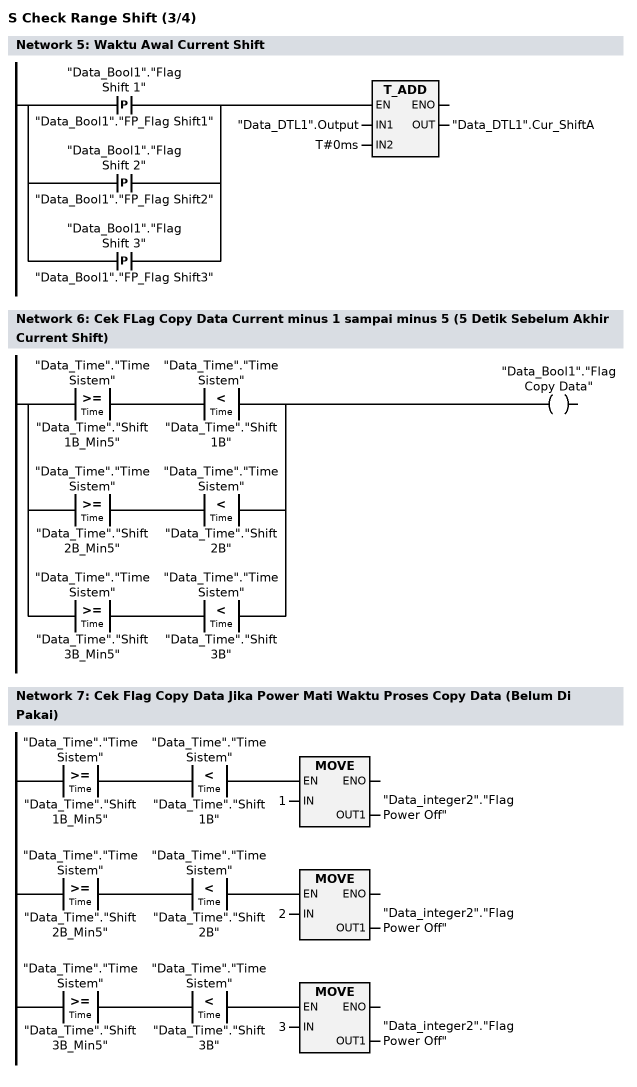
   #_w1 := "Data_Bool1"."Flag Shift 1" AND NOT "Data_Bool1"."FP_Flag Shift1";   // rising edge of "Data_Bool1"."Flag Shift 1"
   "Data_Bool1"."FP_Flag Shift1" := "Data_Bool1"."Flag Shift 1";
   #_w2 := "Data_Bool1"."Flag Shift 2" AND NOT "Data_Bool1"."FP_Flag Shift2";   // rising edge of "Data_Bool1"."Flag Shift 2"
   "Data_Bool1"."FP_Flag Shift2" := "Data_Bool1"."Flag Shift 2";
   #_w3 := "Data_Bool1"."Flag Shift 3" AND NOT "Data_Bool1"."FP_Flag Shift3";   // rising edge of "Data_Bool1"."Flag Shift 3"
   "Data_Bool1"."FP_Flag Shift3" := "Data_Bool1"."Flag Shift 3";
   IF #_w1 OR #_w2 OR #_w3 THEN
       "Data_DTL1".Cur_ShiftA := T_ADD(IN1 := "Data_DTL1".Output, IN2 := T#0ms);
   END_IF;
END_REGION

REGION Network 6: Cek FLag Copy Data Current minus 1 sampai minus 5 (5 Detik Sebelum Akhir Current Shift)
   RUNG wire#powerrail
      { S7_Templates := "SrcType := Time" } GE_Contact(in1 := "Data_Time"."Time Sistem", in2 := "Data_Time"."Shift 1B_Min5")
      { S7_Templates := "SrcType := Time" } LT_Contact(in1 := "Data_Time"."Time Sistem", in2 := "Data_Time"."Shift 1B")
      wire#w1
      Coil( "Data_Bool1"."Flag Copy Data" )
   END_RUNG
   RUNG wire#powerrail
      { S7_Templates := "SrcType := Time" } GE_Contact(in1 := "Data_Time"."Time Sistem", in2 := "Data_Time"."Shift 2B_Min5")
      { S7_Templates := "SrcType := Time" } LT_Contact(in1 := "Data_Time"."Time Sistem", in2 := "Data_Time"."Shift 2B")
   END_RUNG wire#w1
   RUNG wire#powerrail
      { S7_Templates := "SrcType := Time" } GE_Contact(in1 := "Data_Time"."Time Sistem", in2 := "Data_Time"."Shift 3B_Min5")
      { S7_Templates := "SrcType := Time" } LT_Contact(in1 := "Data_Time"."Time Sistem", in2 := "Data_Time"."Shift 3B")
   END_RUNG wire#w1
   // the same network as SCL:
   "Data_Bool1"."Flag Copy Data" := (("Data_Time"."Time Sistem" >= "Data_Time"."Shift 1B_Min5") AND ("Data_Time"."Time Sistem" < "Data_Time"."Shift 1B")) OR (("Data_Time"."Time Sistem" >= "Data_Time"."Shift 2B_Min5") AND ("Data_Time"."Time Sistem" < "Data_Time"."Shift 2B")) OR (("Data_Time"."Time Sistem" >= "Data_Time"."Shift 3B_Min5") AND ("Data_Time"."Time Sistem" < "Data_Time"."Shift 3B"));
END_REGION

REGION Network 7: Cek Flag Copy Data Jika Power Mati Waktu Proses Copy Data (Belum Di Pakai)
   RUNG wire#powerrail
      { S7_Templates := "SrcType := Time" } GE_Contact(in1 := "Data_Time"."Time Sistem", in2 := "Data_Time"."Shift 1B_Min5")
      { S7_Templates := "SrcType := Time" } LT_Contact(in1 := "Data_Time"."Time Sistem", in2 := "Data_Time"."Shift 1B")
      { S7_GenerateENO := "TRUE" } Move(in := 1, out1 => "Data_integer2"."Flag Power Off")
   END_RUNG
   RUNG wire#powerrail
      { S7_Templates := "SrcType := Time" } GE_Contact(in1 := "Data_Time"."Time Sistem", in2 := "Data_Time"."Shift 2B_Min5")
      { S7_Templates := "SrcType := Time" } LT_Contact(in1 := "Data_Time"."Time Sistem", in2 := "Data_Time"."Shift 2B")
      { S7_GenerateENO := "TRUE" } Move(in := 2, out1 => "Data_integer2"."Flag Power Off")
   END_RUNG
   RUNG wire#powerrail
      { S7_Templates := "SrcType := Time" } GE_Contact(in1 := "Data_Time"."Time Sistem", in2 := "Data_Time"."Shift 3B_Min5")
      { S7_Templates := "SrcType := Time" } LT_Contact(in1 := "Data_Time"."Time Sistem", in2 := "Data_Time"."Shift 3B")
      { S7_GenerateENO := "TRUE" } Move(in := 3, out1 => "Data_integer2"."Flag Power Off")
   END_RUNG
   // the same network as SCL:
   IF ("Data_Time"."Time Sistem" >= "Data_Time"."Shift 1B_Min5") AND ("Data_Time"."Time Sistem" < "Data_Time"."Shift 1B") THEN
       "Data_integer2"."Flag Power Off" := 1;
   END_IF;
   IF ("Data_Time"."Time Sistem" >= "Data_Time"."Shift 2B_Min5") AND ("Data_Time"."Time Sistem" < "Data_Time"."Shift 2B") THEN
       "Data_integer2"."Flag Power Off" := 2;
   END_IF;
   IF ("Data_Time"."Time Sistem" >= "Data_Time"."Shift 3B_Min5") AND ("Data_Time"."Time Sistem" < "Data_Time"."Shift 3B") THEN
       "Data_integer2"."Flag Power Off" := 3;
   END_IF;
END_REGION

REGION Network 8: Waktu Awal Current Shift Static Dan Set Copi data Setelah Power mati di waktu proses Copi Data (belum Dipakai)
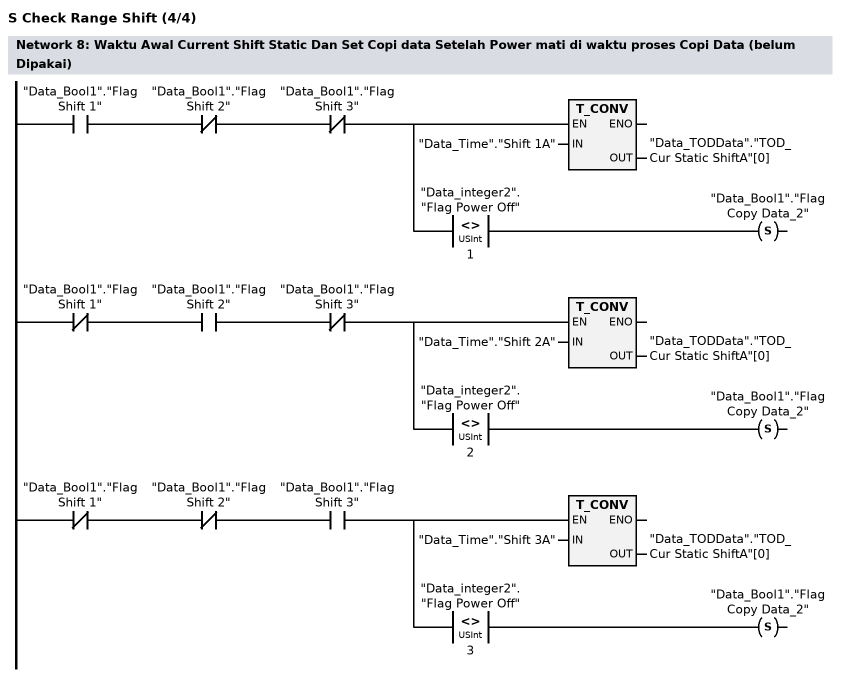
   #_w1 := "Data_Bool1"."Flag Shift 1" AND NOT "Data_Bool1"."Flag Shift 2" AND NOT "Data_Bool1"."Flag Shift 3";
   IF #_w1 THEN "Data_TODData"."TOD_Cur Static ShiftA"[0] := T_CONV(IN := "Data_Time"."Shift 1A"); END_IF;
   IF #_w1 AND ("Data_integer2"."Flag Power Off" <> 1) THEN "Data_Bool1"."Flag Copy Data_2" := TRUE; END_IF;
   #_w2 := NOT "Data_Bool1"."Flag Shift 1" AND "Data_Bool1"."Flag Shift 2" AND NOT "Data_Bool1"."Flag Shift 3";
   IF #_w2 THEN "Data_TODData"."TOD_Cur Static ShiftA"[0] := T_CONV(IN := "Data_Time"."Shift 2A"); END_IF;
   IF #_w2 AND ("Data_integer2"."Flag Power Off" <> 2) THEN "Data_Bool1"."Flag Copy Data_2" := TRUE; END_IF;
   #_w3 := NOT "Data_Bool1"."Flag Shift 1" AND NOT "Data_Bool1"."Flag Shift 2" AND "Data_Bool1"."Flag Shift 3";
   IF #_w3 THEN "Data_TODData"."TOD_Cur Static ShiftA"[0] := T_CONV(IN := "Data_Time"."Shift 3A"); END_IF;
   IF #_w3 AND ("Data_integer2"."Flag Power Off" <> 3) THEN "Data_Bool1"."Flag Copy Data_2" := TRUE; END_IF;
END_REGION
END_FUNCTION_BLOCK

FUNCTION_BLOCK "S Block Current Shift_M2"   // FB11, LAD
{ S7_Optimized_Access := 'TRUE' }
VERSION : 0.1
BEGIN

REGION Network 1: Move Date Time M2
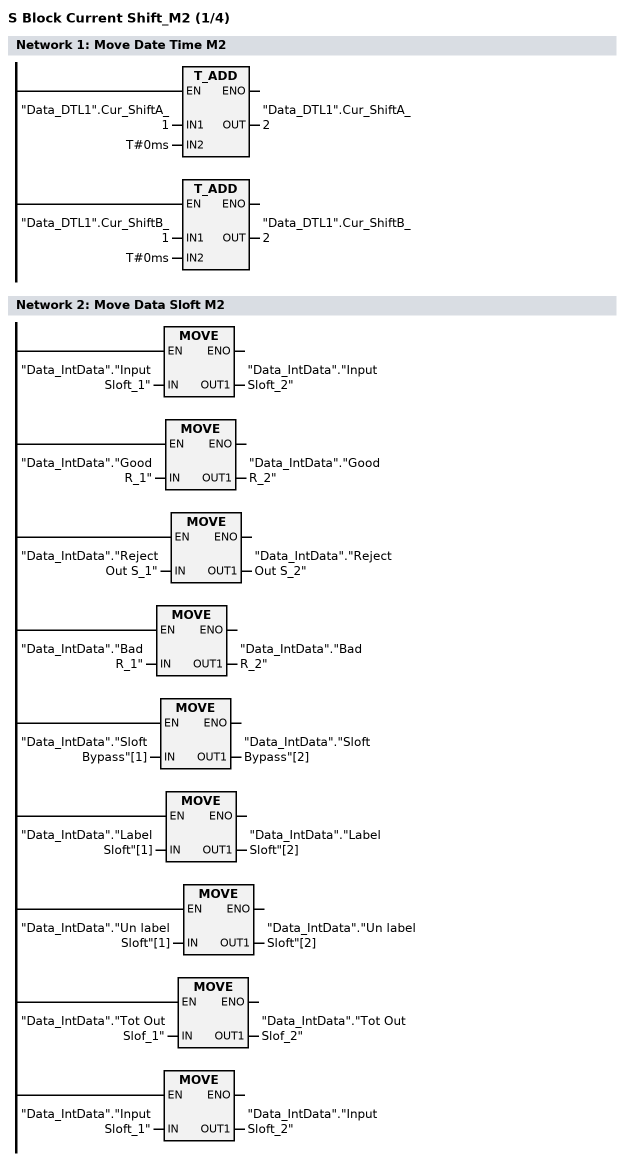
   "Data_DTL1".Cur_ShiftA_2 := T_ADD(IN1 := "Data_DTL1".Cur_ShiftA_1, IN2 := T#0ms);
   "Data_DTL1".Cur_ShiftB_2 := T_ADD(IN1 := "Data_DTL1".Cur_ShiftB_1, IN2 := T#0ms);
END_REGION

REGION Network 2: Move Data Sloft M2
   RUNG wire#powerrail
      { S7_GenerateENO := "TRUE" } Move(in := "Data_IntData"."Input Sloft_1", out1 => "Data_IntData"."Input Sloft_2")
   END_RUNG
   RUNG wire#powerrail
      { S7_GenerateENO := "TRUE" } Move(in := "Data_IntData"."Good R_1", out1 => "Data_IntData"."Good R_2")
   END_RUNG
   RUNG wire#powerrail
      { S7_GenerateENO := "TRUE" } Move(in := "Data_IntData"."Reject Out S_1", out1 => "Data_IntData"."Reject Out S_2")
   END_RUNG
   RUNG wire#powerrail
      { S7_GenerateENO := "TRUE" } Move(in := "Data_IntData"."Bad R_1", out1 => "Data_IntData"."Bad R_2")
   END_RUNG
   RUNG wire#powerrail
      { S7_GenerateENO := "TRUE" } Move(in := "Data_IntData"."Sloft Bypass"[1], out1 => "Data_IntData"."Sloft Bypass"[2])
   END_RUNG
   RUNG wire#powerrail
      { S7_GenerateENO := "TRUE" } Move(in := "Data_IntData"."Label Sloft"[1], out1 => "Data_IntData"."Label Sloft"[2])
   END_RUNG
   RUNG wire#powerrail
      { S7_GenerateENO := "TRUE" } Move(in := "Data_IntData"."Un label Sloft"[1], out1 => "Data_IntData"."Un label Sloft"[2])
   END_RUNG
   RUNG wire#powerrail
      { S7_GenerateENO := "TRUE" } Move(in := "Data_IntData"."Tot Out Slof_1", out1 => "Data_IntData"."Tot Out Slof_2")
   END_RUNG
   RUNG wire#powerrail
      { S7_GenerateENO := "TRUE" } Move(in := "Data_IntData"."Input Sloft_1", out1 => "Data_IntData"."Input Sloft_2")
   END_RUNG
   // the same network as SCL:
   "Data_IntData"."Input Sloft_2" := "Data_IntData"."Input Sloft_1";
   "Data_IntData"."Good R_2" := "Data_IntData"."Good R_1";
   "Data_IntData"."Reject Out S_2" := "Data_IntData"."Reject Out S_1";
   "Data_IntData"."Bad R_2" := "Data_IntData"."Bad R_1";
   "Data_IntData"."Sloft Bypass"[2] := "Data_IntData"."Sloft Bypass"[1];
   "Data_IntData"."Label Sloft"[2] := "Data_IntData"."Label Sloft"[1];
   "Data_IntData"."Un label Sloft"[2] := "Data_IntData"."Un label Sloft"[1];
   "Data_IntData"."Tot Out Slof_2" := "Data_IntData"."Tot Out Slof_1";
   "Data_IntData"."Input Sloft_2" := "Data_IntData"."Input Sloft_1";
END_REGION

REGION Network 3: Move Data Sloft Trigger & Aplicator M2
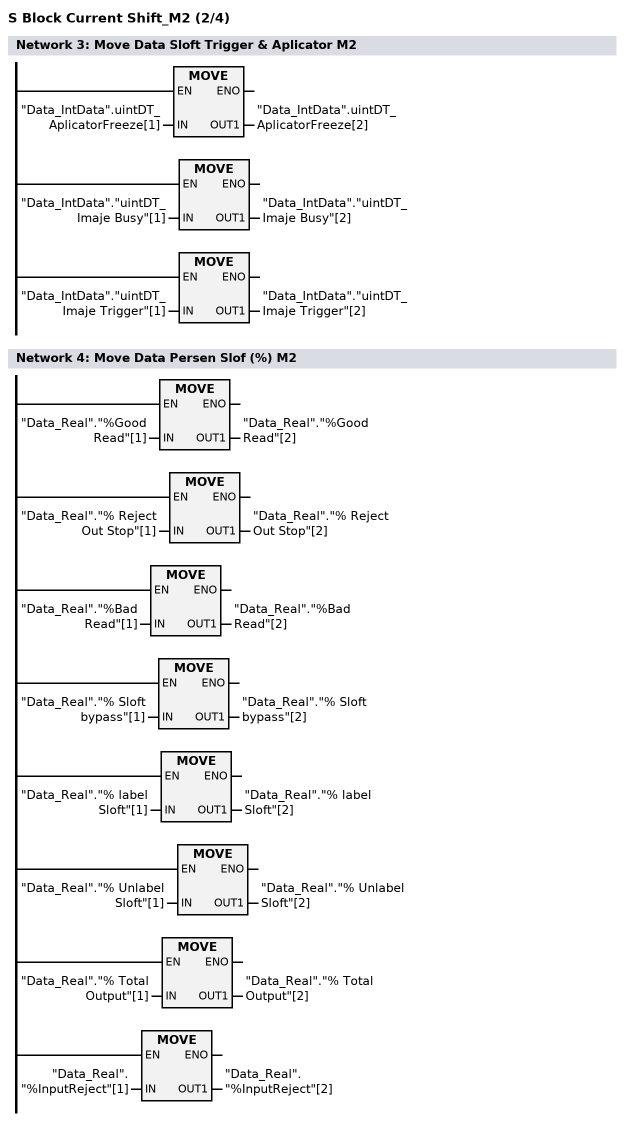
   RUNG wire#powerrail
      { S7_GenerateENO := "TRUE" } Move(in := "Data_IntData".uintDT_AplicatorFreeze[1], out1 => "Data_IntData".uintDT_AplicatorFreeze[2])
   END_RUNG
   RUNG wire#powerrail
      { S7_GenerateENO := "TRUE" } Move(in := "Data_IntData"."uintDT_Imaje Busy"[1], out1 => "Data_IntData"."uintDT_Imaje Busy"[2])
   END_RUNG
   RUNG wire#powerrail
      { S7_GenerateENO := "TRUE" } Move(in := "Data_IntData"."uintDT_Imaje Trigger"[1], out1 => "Data_IntData"."uintDT_Imaje Trigger"[2])
   END_RUNG
   // the same network as SCL:
   "Data_IntData".uintDT_AplicatorFreeze[2] := "Data_IntData".uintDT_AplicatorFreeze[1];
   "Data_IntData"."uintDT_Imaje Busy"[2] := "Data_IntData"."uintDT_Imaje Busy"[1];
   "Data_IntData"."uintDT_Imaje Trigger"[2] := "Data_IntData"."uintDT_Imaje Trigger"[1];
END_REGION

REGION Network 4: Move Data Persen Slof (%) M2
   RUNG wire#powerrail
      { S7_GenerateENO := "TRUE" } Move(in := "Data_Real"."%Good Read"[1], out1 => "Data_Real"."%Good Read"[2])
   END_RUNG
   RUNG wire#powerrail
      { S7_GenerateENO := "TRUE" } Move(in := "Data_Real"."% Reject Out Stop"[1], out1 => "Data_Real"."% Reject Out Stop"[2])
   END_RUNG
   RUNG wire#powerrail
      { S7_GenerateENO := "TRUE" } Move(in := "Data_Real"."%Bad Read"[1], out1 => "Data_Real"."%Bad Read"[2])
   END_RUNG
   RUNG wire#powerrail
      { S7_GenerateENO := "TRUE" } Move(in := "Data_Real"."% Sloft bypass"[1], out1 => "Data_Real"."% Sloft bypass"[2])
   END_RUNG
   RUNG wire#powerrail
      { S7_GenerateENO := "TRUE" } Move(in := "Data_Real"."% label Sloft"[1], out1 => "Data_Real"."% label Sloft"[2])
   END_RUNG
   RUNG wire#powerrail
      { S7_GenerateENO := "TRUE" } Move(in := "Data_Real"."% Unlabel Sloft"[1], out1 => "Data_Real"."% Unlabel Sloft"[2])
   END_RUNG
   RUNG wire#powerrail
      { S7_GenerateENO := "TRUE" } Move(in := "Data_Real"."% Total Output"[1], out1 => "Data_Real"."% Total Output"[2])
   END_RUNG
   RUNG wire#powerrail
      { S7_GenerateENO := "TRUE" } Move(in := "Data_Real"."%InputReject"[1], out1 => "Data_Real"."%InputReject"[2])
   END_RUNG
   // the same network as SCL:
   "Data_Real"."%Good Read"[2] := "Data_Real"."%Good Read"[1];
   "Data_Real"."% Reject Out Stop"[2] := "Data_Real"."% Reject Out Stop"[1];
   "Data_Real"."%Bad Read"[2] := "Data_Real"."%Bad Read"[1];
   "Data_Real"."% Sloft bypass"[2] := "Data_Real"."% Sloft bypass"[1];
   "Data_Real"."% label Sloft"[2] := "Data_Real"."% label Sloft"[1];
   "Data_Real"."% Unlabel Sloft"[2] := "Data_Real"."% Unlabel Sloft"[1];
   "Data_Real"."% Total Output"[2] := "Data_Real"."% Total Output"[1];
   "Data_Real"."%InputReject"[2] := "Data_Real"."%InputReject"[1];
END_REGION

REGION Network 5: Move Data Time Mesin M2
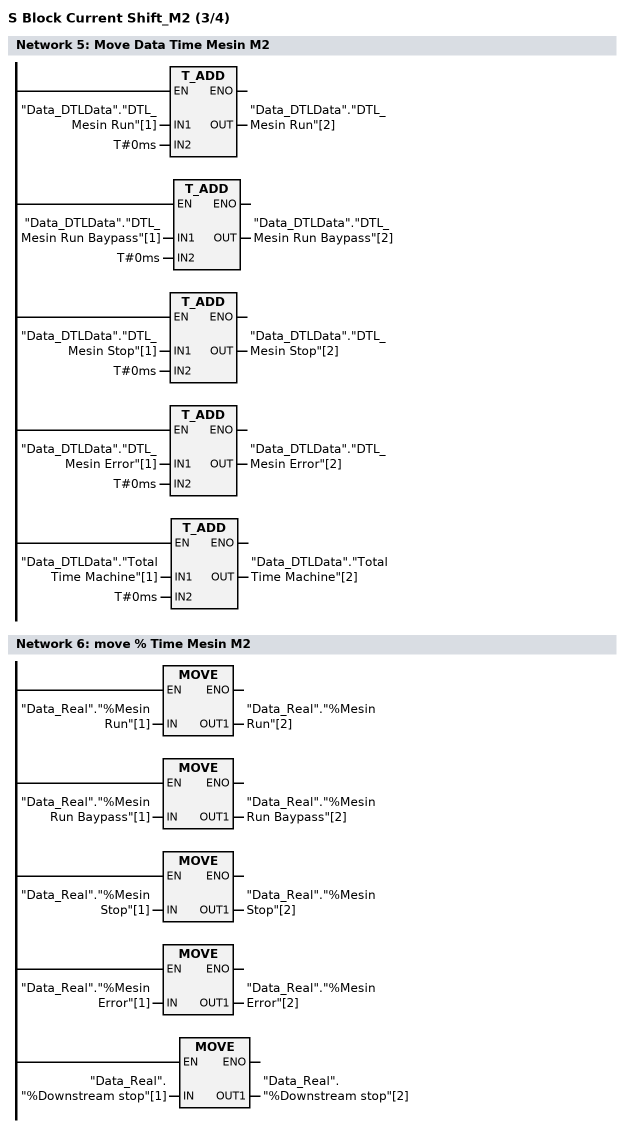
   "Data_DTLData"."DTL_Mesin Run"[2] := T_ADD(IN1 := "Data_DTLData"."DTL_Mesin Run"[1], IN2 := T#0ms);
   "Data_DTLData"."DTL_Mesin Run Baypass"[2] := T_ADD(IN1 := "Data_DTLData"."DTL_Mesin Run Baypass"[1],
                           IN2 := T#0ms);
   "Data_DTLData"."DTL_Mesin Stop"[2] := T_ADD(IN1 := "Data_DTLData"."DTL_Mesin Stop"[1], IN2 := T#0ms);
   "Data_DTLData"."DTL_Mesin Error"[2] := T_ADD(IN1 := "Data_DTLData"."DTL_Mesin Error"[1], IN2 := T#0ms);
   "Data_DTLData"."Total Time Machine"[2] := T_ADD(IN1 := "Data_DTLData"."Total Time Machine"[1], IN2 := T#0ms);
END_REGION

REGION Network 6: move % Time Mesin M2
   RUNG wire#powerrail
      { S7_GenerateENO := "TRUE" } Move(in := "Data_Real"."%Mesin Run"[1], out1 => "Data_Real"."%Mesin Run"[2])
   END_RUNG
   RUNG wire#powerrail
      { S7_GenerateENO := "TRUE" } Move(in := "Data_Real"."%Mesin Run Baypass"[1], out1 => "Data_Real"."%Mesin Run Baypass"[2])
   END_RUNG
   RUNG wire#powerrail
      { S7_GenerateENO := "TRUE" } Move(in := "Data_Real"."%Mesin Stop"[1], out1 => "Data_Real"."%Mesin Stop"[2])
   END_RUNG
   RUNG wire#powerrail
      { S7_GenerateENO := "TRUE" } Move(in := "Data_Real"."%Mesin Error"[1], out1 => "Data_Real"."%Mesin Error"[2])
   END_RUNG
   RUNG wire#powerrail
      { S7_GenerateENO := "TRUE" } Move(in := "Data_Real"."%Downstream stop"[1], out1 => "Data_Real"."%Downstream stop"[2])
   END_RUNG
   // the same network as SCL:
   "Data_Real"."%Mesin Run"[2] := "Data_Real"."%Mesin Run"[1];
   "Data_Real"."%Mesin Run Baypass"[2] := "Data_Real"."%Mesin Run Baypass"[1];
   "Data_Real"."%Mesin Stop"[2] := "Data_Real"."%Mesin Stop"[1];
   "Data_Real"."%Mesin Error"[2] := "Data_Real"."%Mesin Error"[1];
   "Data_Real"."%Downstream stop"[2] := "Data_Real"."%Downstream stop"[1];
END_REGION

REGION Network 7: Move Counter Error M2
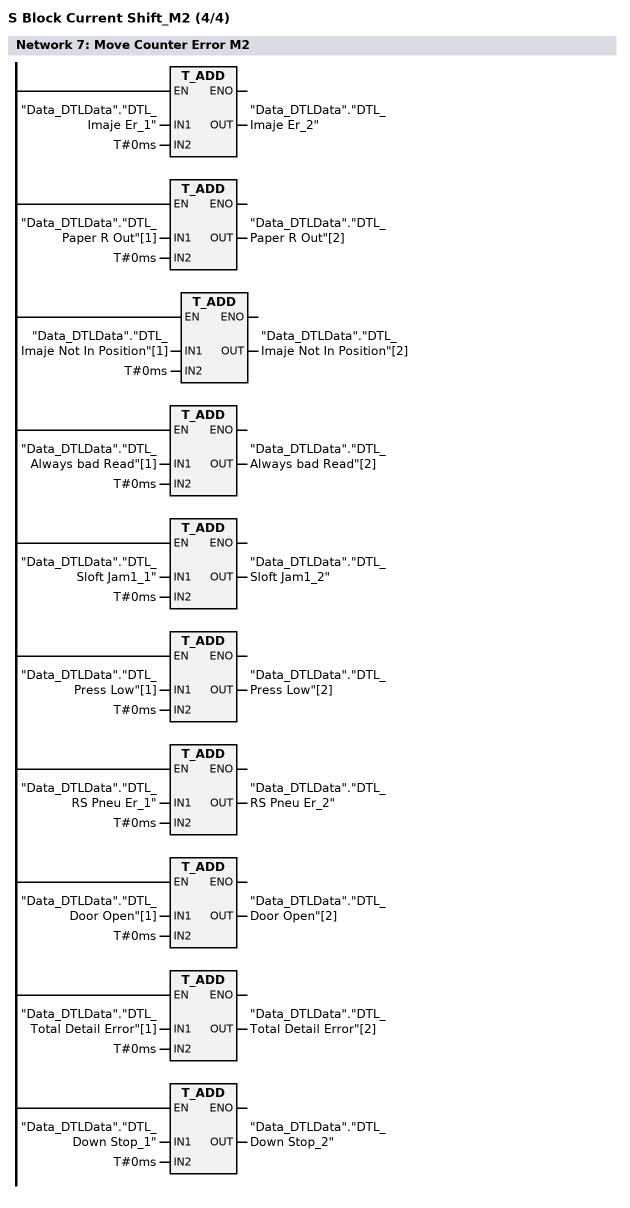
   "Data_DTLData"."DTL_Imaje Er_2" := T_ADD(IN1 := "Data_DTLData"."DTL_Imaje Er_1", IN2 := T#0ms);
   "Data_DTLData"."DTL_Paper R Out"[2] := T_ADD(IN1 := "Data_DTLData"."DTL_Paper R Out"[1], IN2 := T#0ms);
   "Data_DTLData"."DTL_Imaje Not In Position"[2] := T_ADD(IN1 := "Data_DTLData"."DTL_Imaje Not In Position"[1],
                           IN2 := T#0ms);
   "Data_DTLData"."DTL_Always bad Read"[2] := T_ADD(IN1 := "Data_DTLData"."DTL_Always bad Read"[1],
                           IN2 := T#0ms);
   "Data_DTLData"."DTL_Sloft Jam1_2" := T_ADD(IN1 := "Data_DTLData"."DTL_Sloft Jam1_1", IN2 := T#0ms);
   "Data_DTLData"."DTL_Press Low"[2] := T_ADD(IN1 := "Data_DTLData"."DTL_Press Low"[1], IN2 := T#0ms);
   "Data_DTLData"."DTL_RS Pneu Er_2" := T_ADD(IN1 := "Data_DTLData"."DTL_RS Pneu Er_1", IN2 := T#0ms);
   "Data_DTLData"."DTL_Door Open"[2] := T_ADD(IN1 := "Data_DTLData"."DTL_Door Open"[1], IN2 := T#0ms);
   "Data_DTLData"."DTL_Total Detail Error"[2] := T_ADD(IN1 := "Data_DTLData"."DTL_Total Detail Error"[1],
                           IN2 := T#0ms);
   "Data_DTLData"."DTL_Down Stop_2" := T_ADD(IN1 := "Data_DTLData"."DTL_Down Stop_1", IN2 := T#0ms);
END_REGION
END_FUNCTION_BLOCK

FUNCTION_BLOCK "S Block Current Shift_M3"   // FB12, LAD
{ S7_Optimized_Access := 'TRUE' }
VERSION : 0.1
BEGIN

REGION Network 1: Move Date Time M3